(* Logix 5000 project; controller PLC_MCC1201_220AP1 vendor 1 type 14 code 164 rev 35.11; software revision 35.00; part 6 of 25 *)
(* tags used below, declared in another part *)
   B3 : DINT[102];
   HMI_Alarm_Reset : BOOL;   // HMI_Alarm_Reset
   HMI_MAN_CMD_WR : UDT_MAN_CMD_WR;
   LEHR_SPEED : ALIAS FOR N60[1];
   M206_M1_DR : AXIS_CIP_DRIVE;
   M207_M1_DR : AXIS_CIP_DRIVE;
   M208_M1_DR : AXIS_CIP_DRIVE;
   M209_M1_DR : AXIS_CIP_DRIVE;
   M2xx_CONVEYOR : MAC_CONVEYOR[20];
   M2xx_CONVEYOR_IN_MOTION : MAC_CONVEYOR_IN_MOTION[20];
   M2xx_CONVEYOR_OUT_MOTION : MAC_CONVEYOR_OUT_MOTION[20];
   TMP_dDirection : DINT;
   TMP_rAcc : REAL;
   TMP_rDec : REAL;
   TMP_rSpeed : REAL;
   TMP_xAlwaysOFF : BOOL;
   TMP_xRun : BOOL;
(* CommandLogic, continued *)

ROUTINE M206_Conveyor_Motion_Output   (* ladder *)
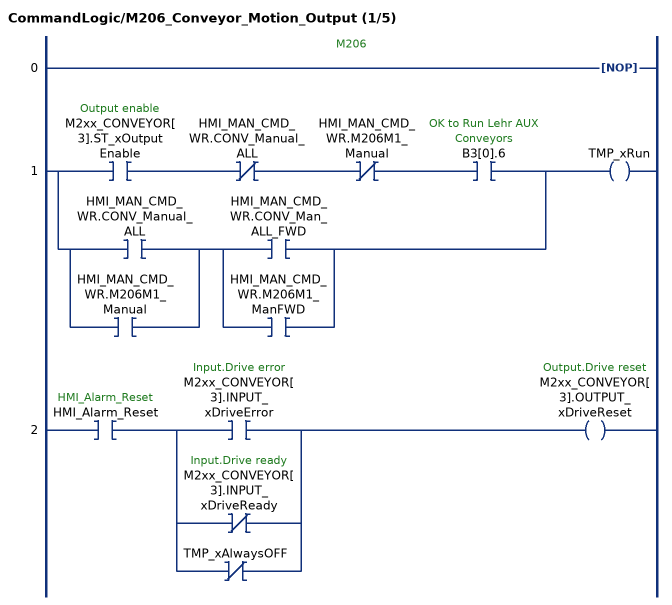
   // M206
   0: NOP();
   1: [XIC(M2xx_CONVEYOR[3].ST_xOutputEnable) XIO(HMI_MAN_CMD_WR.CONV_Manual_ALL) XIO(HMI_MAN_CMD_WR.M206M1_Manual) XIC(B3[0].6) ,[XIC(HMI_MAN_CMD_WR.CONV_Manual_ALL) ,XIC(HMI_MAN_CMD_WR.M206M1_Manual) ] [XIC(HMI_MAN_CMD_WR.CONV_Man_ALL_FWD) ,XIC(HMI_MAN_CMD_WR.M206M1_ManFWD) ] ]OTE(TMP_xRun);
   2: XIC(HMI_Alarm_Reset)[XIC(M2xx_CONVEYOR[3].INPUT_xDriveError) ,XIO(M2xx_CONVEYOR[3].INPUT_xDriveReady) ,XIO(TMP_xAlwaysOFF) ]OTE(M2xx_CONVEYOR[3].OUTPUT_xDriveReset);
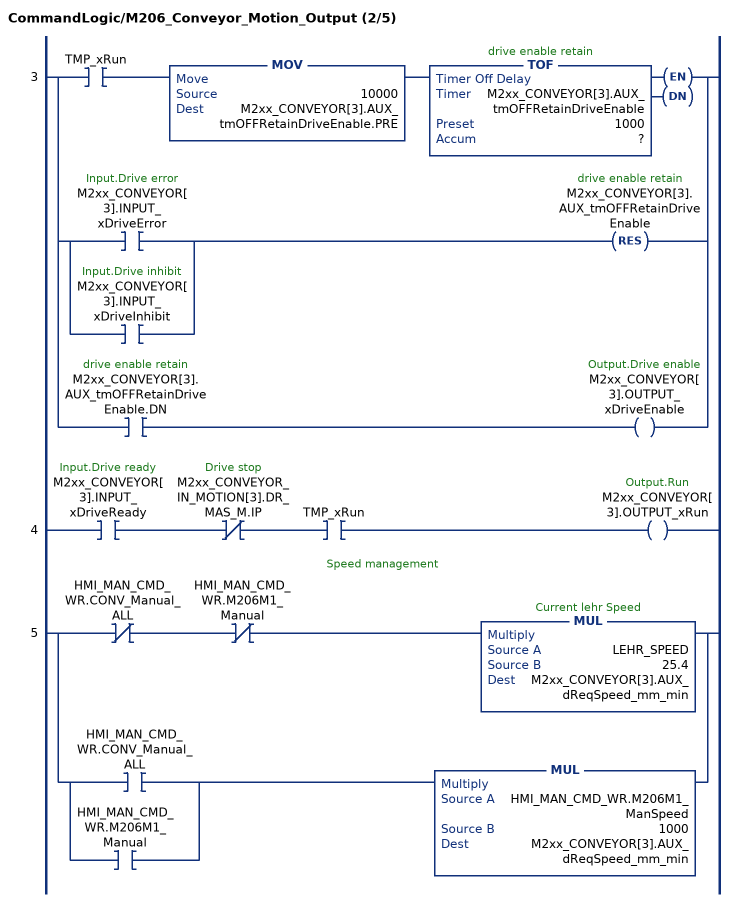
   3: [XIC(TMP_xRun) MOV(10000,M2xx_CONVEYOR[3].AUX_tmOFFRetainDriveEnable.PRE) TOF(M2xx_CONVEYOR[3].AUX_tmOFFRetainDriveEnable,?,?) ,[XIC(M2xx_CONVEYOR[3].INPUT_xDriveError) ,XIC(M2xx_CONVEYOR[3].INPUT_xDriveInhibit) ] RES(M2xx_CONVEYOR[3].AUX_tmOFFRetainDriveEnable) ,XIC(M2xx_CONVEYOR[3].AUX_tmOFFRetainDriveEnable.DN) OTE(M2xx_CONVEYOR[3].OUTPUT_xDriveEnable) ];
   4: XIC(M2xx_CONVEYOR[3].INPUT_xDriveReady)XIO(M2xx_CONVEYOR_IN_MOTION[3].DR_MAS_M.IP)XIC(TMP_xRun)OTE(M2xx_CONVEYOR[3].OUTPUT_xRun);
   // Speed management
   5: [XIO(HMI_MAN_CMD_WR.CONV_Manual_ALL) XIO(HMI_MAN_CMD_WR.M206M1_Manual) MUL(LEHR_SPEED,25.4,M2xx_CONVEYOR[3].AUX_dReqSpeed_mm_min) ,[XIC(HMI_MAN_CMD_WR.CONV_Manual_ALL) ,XIC(HMI_MAN_CMD_WR.M206M1_Manual) ] MUL(HMI_MAN_CMD_WR.M206M1_ManSpeed,1000,M2xx_CONVEYOR[3].AUX_dReqSpeed_mm_min) ];
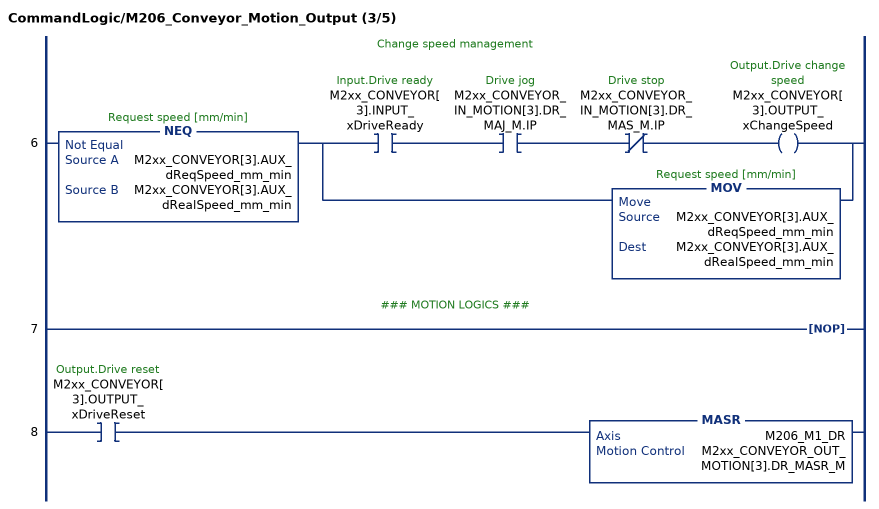
   // Change speed management
   6: NEQ(M2xx_CONVEYOR[3].AUX_dReqSpeed_mm_min,M2xx_CONVEYOR[3].AUX_dRealSpeed_mm_min)[XIC(M2xx_CONVEYOR[3].INPUT_xDriveReady) XIC(M2xx_CONVEYOR_IN_MOTION[3].DR_MAJ_M.IP) XIO(M2xx_CONVEYOR_IN_MOTION[3].DR_MAS_M.IP) OTE(M2xx_CONVEYOR[3].OUTPUT_xChangeSpeed) ,MOV(M2xx_CONVEYOR[3].AUX_dReqSpeed_mm_min,M2xx_CONVEYOR[3].AUX_dRealSpeed_mm_min) ];
   // ### MOTION LOGICS ###
   7: NOP();
   8: XIC(M2xx_CONVEYOR[3].OUTPUT_xDriveReset)MASR(M206_M1_DR,M2xx_CONVEYOR_OUT_MOTION[3].DR_MASR_M);
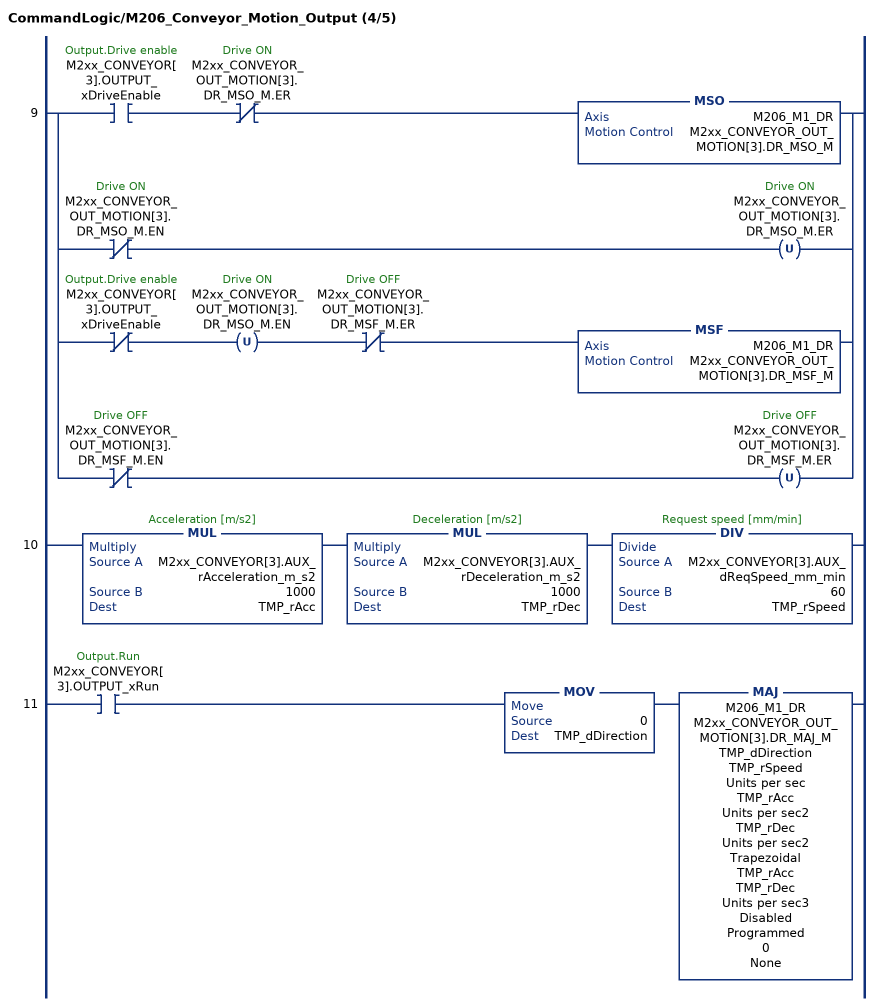
   9: [XIC(M2xx_CONVEYOR[3].OUTPUT_xDriveEnable) XIO(M2xx_CONVEYOR_OUT_MOTION[3].DR_MSO_M.ER) MSO(M206_M1_DR,M2xx_CONVEYOR_OUT_MOTION[3].DR_MSO_M) ,XIO(M2xx_CONVEYOR_OUT_MOTION[3].DR_MSO_M.EN) OTU(M2xx_CONVEYOR_OUT_MOTION[3].DR_MSO_M.ER) ,XIO(M2xx_CONVEYOR[3].OUTPUT_xDriveEnable) OTU(M2xx_CONVEYOR_OUT_MOTION[3].DR_MSO_M.EN) XIO(M2xx_CONVEYOR_OUT_MOTION[3].DR_MSF_M.ER) MSF(M206_M1_DR,M2xx_CONVEYOR_OUT_MOTION[3].DR_MSF_M) ,XIO(M2xx_CONVEYOR_OUT_MOTION[3].DR_MSF_M.EN) OTU(M2xx_CONVEYOR_OUT_MOTION[3].DR_MSF_M.ER) ];
   10: MUL(M2xx_CONVEYOR[3].AUX_rAcceleration_m_s2,1000,TMP_rAcc)MUL(M2xx_CONVEYOR[3].AUX_rDeceleration_m_s2,1000,TMP_rDec)DIV(M2xx_CONVEYOR[3].AUX_dReqSpeed_mm_min,60,TMP_rSpeed);
   11: XIC(M2xx_CONVEYOR[3].OUTPUT_xRun)MOV(0,TMP_dDirection)MAJ(M206_M1_DR,M2xx_CONVEYOR_OUT_MOTION[3].DR_MAJ_M,TMP_dDirection,TMP_rSpeed,Units per sec,TMP_rAcc,Units per sec2,TMP_rDec,Units per sec2,Trapezoidal,TMP_rAcc,TMP_rDec,Units per sec3,Disabled,Programmed,0,None);
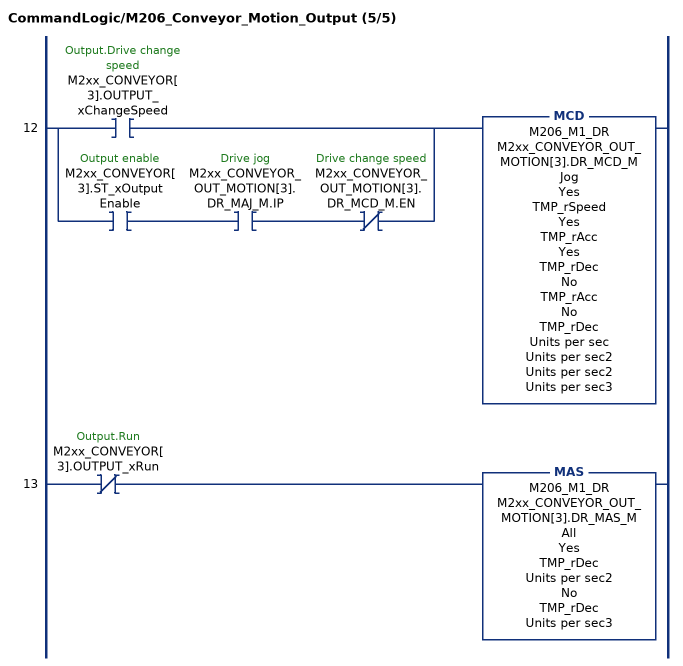
   12: [XIC(M2xx_CONVEYOR[3].OUTPUT_xChangeSpeed) ,XIC(M2xx_CONVEYOR[3].ST_xOutputEnable) XIC(M2xx_CONVEYOR_OUT_MOTION[3].DR_MAJ_M.IP) XIO(M2xx_CONVEYOR_OUT_MOTION[3].DR_MCD_M.EN) ]MCD(M206_M1_DR,M2xx_CONVEYOR_OUT_MOTION[3].DR_MCD_M,Jog,Yes,TMP_rSpeed,Yes,TMP_rAcc,Yes,TMP_rDec,No,TMP_rAcc,No,TMP_rDec,Units per sec,Units per sec2,Units per sec2,Units per sec3);
   13: XIO(M2xx_CONVEYOR[3].OUTPUT_xRun)MAS(M206_M1_DR,M2xx_CONVEYOR_OUT_MOTION[3].DR_MAS_M,All,Yes,TMP_rDec,Units per sec2,No,TMP_rDec,Units per sec3);
END_ROUTINE

ROUTINE M207_Conveyor_Motion_Output   (* ladder *)
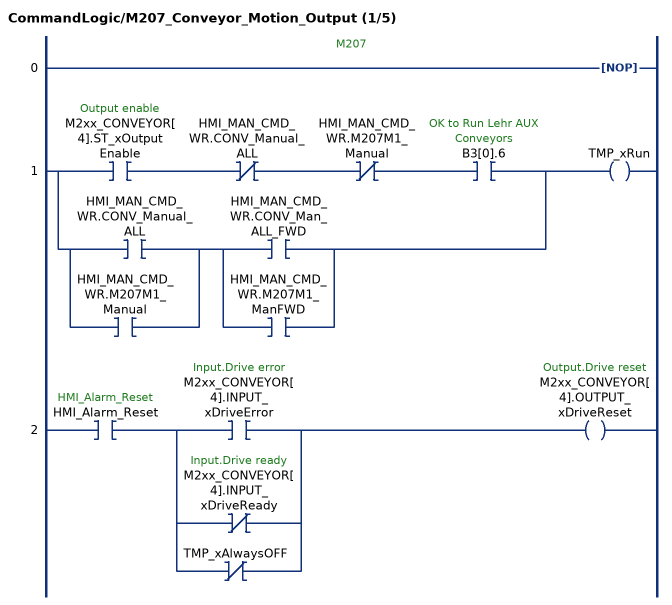
   // M207
   0: NOP();
   1: [XIC(M2xx_CONVEYOR[4].ST_xOutputEnable) XIO(HMI_MAN_CMD_WR.CONV_Manual_ALL) XIO(HMI_MAN_CMD_WR.M207M1_Manual) XIC(B3[0].6) ,[XIC(HMI_MAN_CMD_WR.CONV_Manual_ALL) ,XIC(HMI_MAN_CMD_WR.M207M1_Manual) ] [XIC(HMI_MAN_CMD_WR.CONV_Man_ALL_FWD) ,XIC(HMI_MAN_CMD_WR.M207M1_ManFWD) ] ]OTE(TMP_xRun);
   2: XIC(HMI_Alarm_Reset)[XIC(M2xx_CONVEYOR[4].INPUT_xDriveError) ,XIO(M2xx_CONVEYOR[4].INPUT_xDriveReady) ,XIO(TMP_xAlwaysOFF) ]OTE(M2xx_CONVEYOR[4].OUTPUT_xDriveReset);
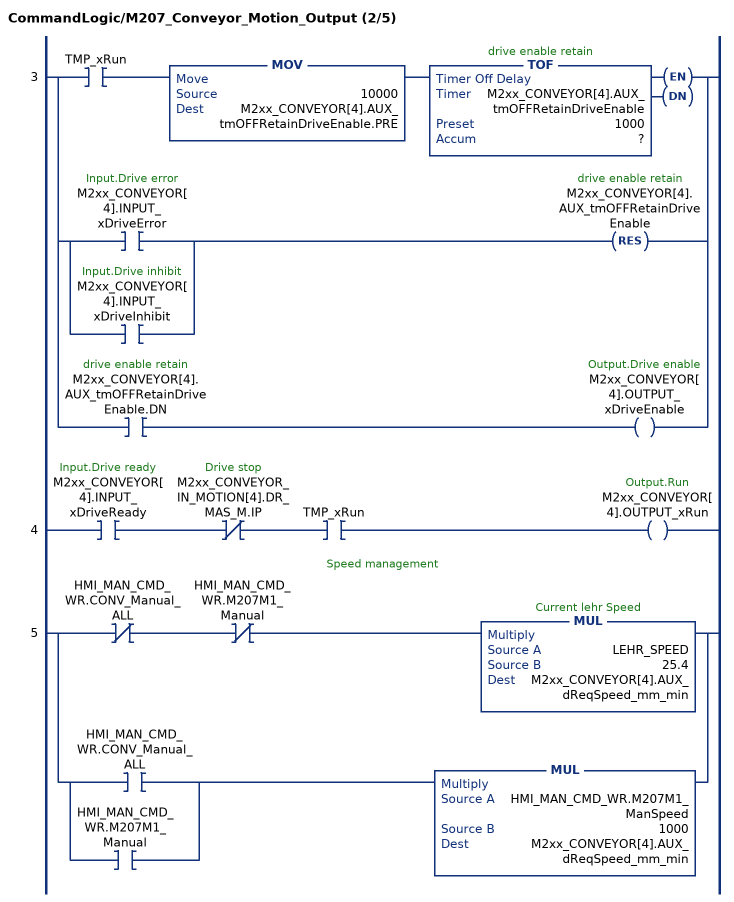
   3: [XIC(TMP_xRun) MOV(10000,M2xx_CONVEYOR[4].AUX_tmOFFRetainDriveEnable.PRE) TOF(M2xx_CONVEYOR[4].AUX_tmOFFRetainDriveEnable,?,?) ,[XIC(M2xx_CONVEYOR[4].INPUT_xDriveError) ,XIC(M2xx_CONVEYOR[4].INPUT_xDriveInhibit) ] RES(M2xx_CONVEYOR[4].AUX_tmOFFRetainDriveEnable) ,XIC(M2xx_CONVEYOR[4].AUX_tmOFFRetainDriveEnable.DN) OTE(M2xx_CONVEYOR[4].OUTPUT_xDriveEnable) ];
   4: XIC(M2xx_CONVEYOR[4].INPUT_xDriveReady)XIO(M2xx_CONVEYOR_IN_MOTION[4].DR_MAS_M.IP)XIC(TMP_xRun)OTE(M2xx_CONVEYOR[4].OUTPUT_xRun);
   // Speed management
   5: [XIO(HMI_MAN_CMD_WR.CONV_Manual_ALL) XIO(HMI_MAN_CMD_WR.M207M1_Manual) MUL(LEHR_SPEED,25.4,M2xx_CONVEYOR[4].AUX_dReqSpeed_mm_min) ,[XIC(HMI_MAN_CMD_WR.CONV_Manual_ALL) ,XIC(HMI_MAN_CMD_WR.M207M1_Manual) ] MUL(HMI_MAN_CMD_WR.M207M1_ManSpeed,1000,M2xx_CONVEYOR[4].AUX_dReqSpeed_mm_min) ];
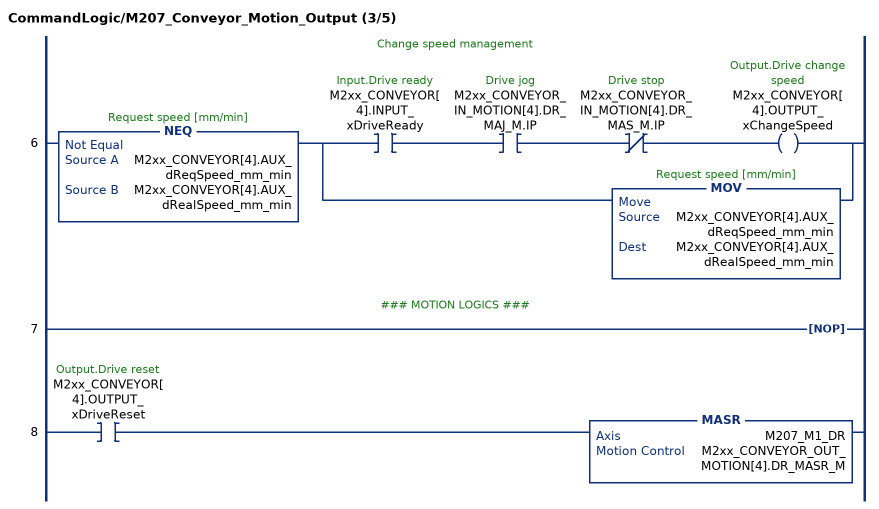
   // Change speed management
   6: NEQ(M2xx_CONVEYOR[4].AUX_dReqSpeed_mm_min,M2xx_CONVEYOR[4].AUX_dRealSpeed_mm_min)[XIC(M2xx_CONVEYOR[4].INPUT_xDriveReady) XIC(M2xx_CONVEYOR_IN_MOTION[4].DR_MAJ_M.IP) XIO(M2xx_CONVEYOR_IN_MOTION[4].DR_MAS_M.IP) OTE(M2xx_CONVEYOR[4].OUTPUT_xChangeSpeed) ,MOV(M2xx_CONVEYOR[4].AUX_dReqSpeed_mm_min,M2xx_CONVEYOR[4].AUX_dRealSpeed_mm_min) ];
   // ### MOTION LOGICS ###
   7: NOP();
   8: XIC(M2xx_CONVEYOR[4].OUTPUT_xDriveReset)MASR(M207_M1_DR,M2xx_CONVEYOR_OUT_MOTION[4].DR_MASR_M);
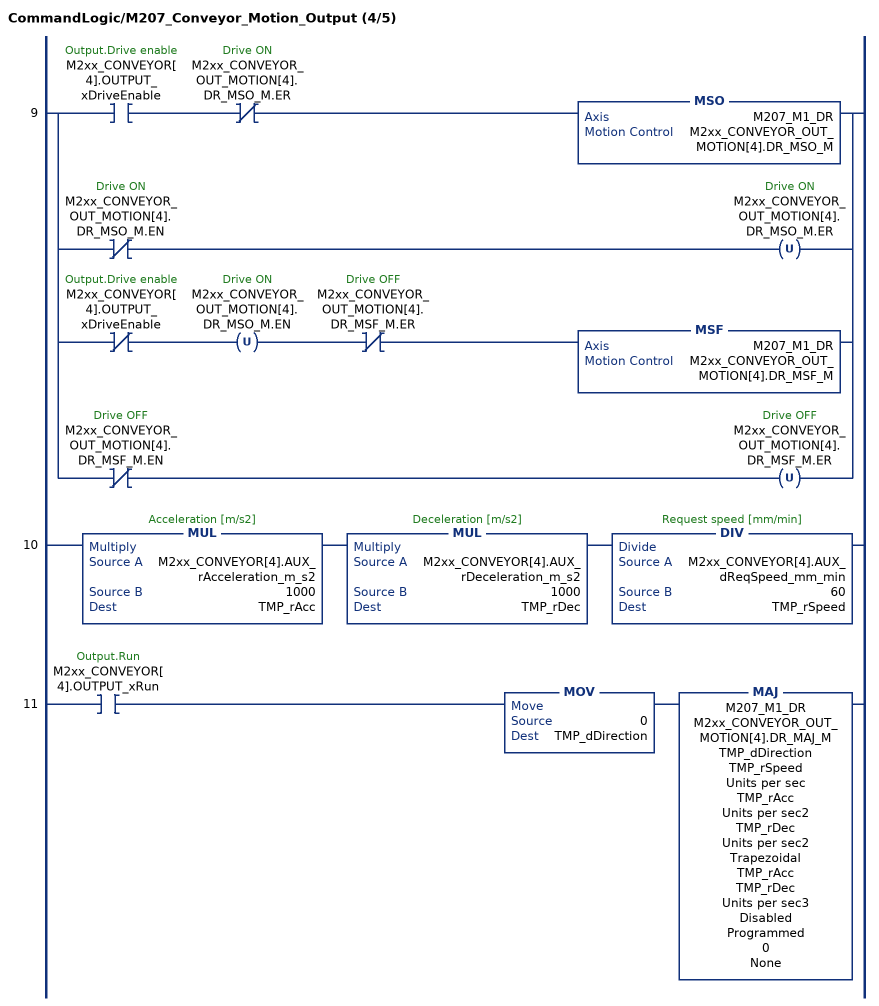
   9: [XIC(M2xx_CONVEYOR[4].OUTPUT_xDriveEnable) XIO(M2xx_CONVEYOR_OUT_MOTION[4].DR_MSO_M.ER) MSO(M207_M1_DR,M2xx_CONVEYOR_OUT_MOTION[4].DR_MSO_M) ,XIO(M2xx_CONVEYOR_OUT_MOTION[4].DR_MSO_M.EN) OTU(M2xx_CONVEYOR_OUT_MOTION[4].DR_MSO_M.ER) ,XIO(M2xx_CONVEYOR[4].OUTPUT_xDriveEnable) OTU(M2xx_CONVEYOR_OUT_MOTION[4].DR_MSO_M.EN) XIO(M2xx_CONVEYOR_OUT_MOTION[4].DR_MSF_M.ER) MSF(M207_M1_DR,M2xx_CONVEYOR_OUT_MOTION[4].DR_MSF_M) ,XIO(M2xx_CONVEYOR_OUT_MOTION[4].DR_MSF_M.EN) OTU(M2xx_CONVEYOR_OUT_MOTION[4].DR_MSF_M.ER) ];
   10: MUL(M2xx_CONVEYOR[4].AUX_rAcceleration_m_s2,1000,TMP_rAcc)MUL(M2xx_CONVEYOR[4].AUX_rDeceleration_m_s2,1000,TMP_rDec)DIV(M2xx_CONVEYOR[4].AUX_dReqSpeed_mm_min,60,TMP_rSpeed);
   11: XIC(M2xx_CONVEYOR[4].OUTPUT_xRun)MOV(0,TMP_dDirection)MAJ(M207_M1_DR,M2xx_CONVEYOR_OUT_MOTION[4].DR_MAJ_M,TMP_dDirection,TMP_rSpeed,Units per sec,TMP_rAcc,Units per sec2,TMP_rDec,Units per sec2,Trapezoidal,TMP_rAcc,TMP_rDec,Units per sec3,Disabled,Programmed,0,None);
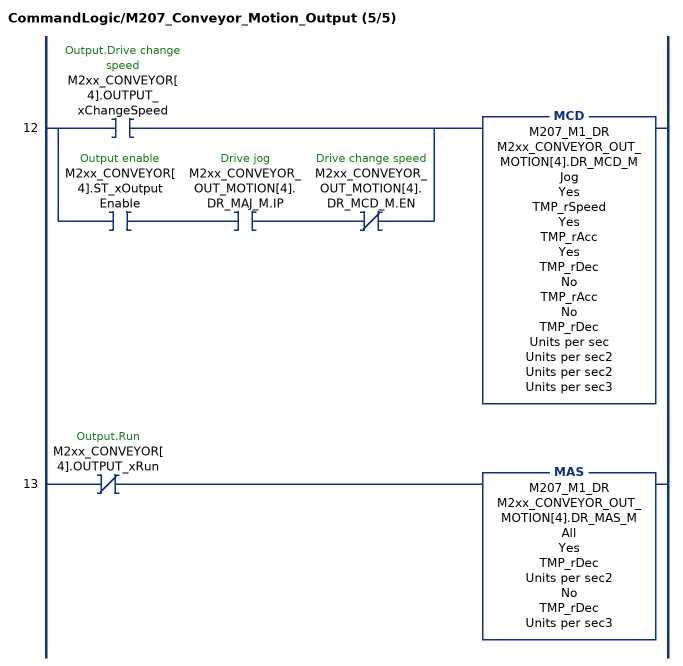
   12: [XIC(M2xx_CONVEYOR[4].OUTPUT_xChangeSpeed) ,XIC(M2xx_CONVEYOR[4].ST_xOutputEnable) XIC(M2xx_CONVEYOR_OUT_MOTION[4].DR_MAJ_M.IP) XIO(M2xx_CONVEYOR_OUT_MOTION[4].DR_MCD_M.EN) ]MCD(M207_M1_DR,M2xx_CONVEYOR_OUT_MOTION[4].DR_MCD_M,Jog,Yes,TMP_rSpeed,Yes,TMP_rAcc,Yes,TMP_rDec,No,TMP_rAcc,No,TMP_rDec,Units per sec,Units per sec2,Units per sec2,Units per sec3);
   13: XIO(M2xx_CONVEYOR[4].OUTPUT_xRun)MAS(M207_M1_DR,M2xx_CONVEYOR_OUT_MOTION[4].DR_MAS_M,All,Yes,TMP_rDec,Units per sec2,No,TMP_rDec,Units per sec3);
END_ROUTINE

ROUTINE M208_Conveyor_Motion_Output   (* ladder *)
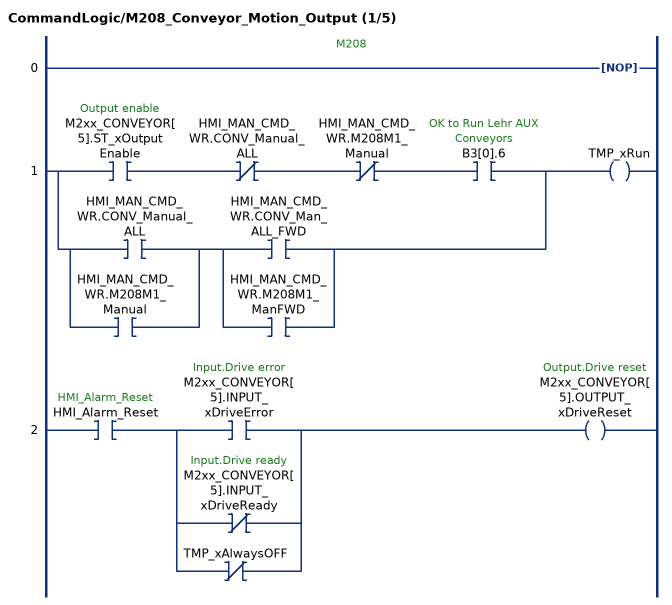
   // M208
   0: NOP();
   1: [XIC(M2xx_CONVEYOR[5].ST_xOutputEnable) XIO(HMI_MAN_CMD_WR.CONV_Manual_ALL) XIO(HMI_MAN_CMD_WR.M208M1_Manual) XIC(B3[0].6) ,[XIC(HMI_MAN_CMD_WR.CONV_Manual_ALL) ,XIC(HMI_MAN_CMD_WR.M208M1_Manual) ] [XIC(HMI_MAN_CMD_WR.CONV_Man_ALL_FWD) ,XIC(HMI_MAN_CMD_WR.M208M1_ManFWD) ] ]OTE(TMP_xRun);
   2: XIC(HMI_Alarm_Reset)[XIC(M2xx_CONVEYOR[5].INPUT_xDriveError) ,XIO(M2xx_CONVEYOR[5].INPUT_xDriveReady) ,XIO(TMP_xAlwaysOFF) ]OTE(M2xx_CONVEYOR[5].OUTPUT_xDriveReset);
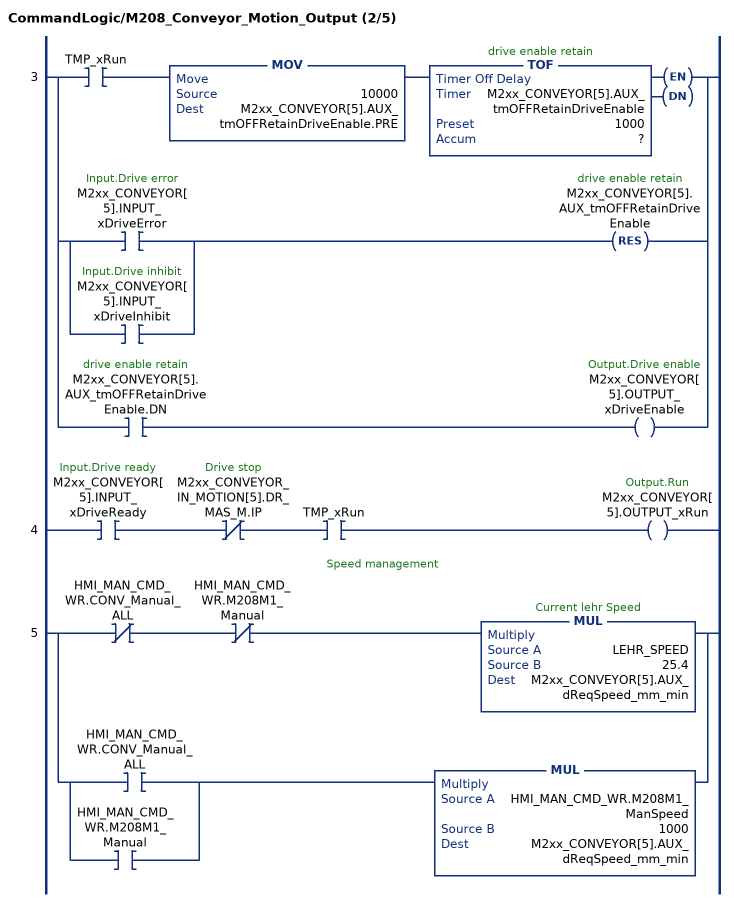
   3: [XIC(TMP_xRun) MOV(10000,M2xx_CONVEYOR[5].AUX_tmOFFRetainDriveEnable.PRE) TOF(M2xx_CONVEYOR[5].AUX_tmOFFRetainDriveEnable,?,?) ,[XIC(M2xx_CONVEYOR[5].INPUT_xDriveError) ,XIC(M2xx_CONVEYOR[5].INPUT_xDriveInhibit) ] RES(M2xx_CONVEYOR[5].AUX_tmOFFRetainDriveEnable) ,XIC(M2xx_CONVEYOR[5].AUX_tmOFFRetainDriveEnable.DN) OTE(M2xx_CONVEYOR[5].OUTPUT_xDriveEnable) ];
   4: XIC(M2xx_CONVEYOR[5].INPUT_xDriveReady)XIO(M2xx_CONVEYOR_IN_MOTION[5].DR_MAS_M.IP)XIC(TMP_xRun)OTE(M2xx_CONVEYOR[5].OUTPUT_xRun);
   // Speed management
   5: [XIO(HMI_MAN_CMD_WR.CONV_Manual_ALL) XIO(HMI_MAN_CMD_WR.M208M1_Manual) MUL(LEHR_SPEED,25.4,M2xx_CONVEYOR[5].AUX_dReqSpeed_mm_min) ,[XIC(HMI_MAN_CMD_WR.CONV_Manual_ALL) ,XIC(HMI_MAN_CMD_WR.M208M1_Manual) ] MUL(HMI_MAN_CMD_WR.M208M1_ManSpeed,1000,M2xx_CONVEYOR[5].AUX_dReqSpeed_mm_min) ];
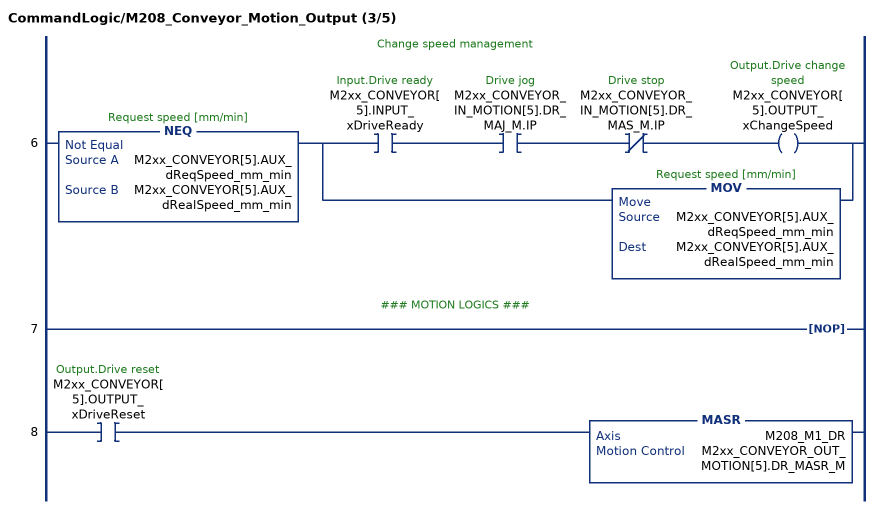
   // Change speed management
   6: NEQ(M2xx_CONVEYOR[5].AUX_dReqSpeed_mm_min,M2xx_CONVEYOR[5].AUX_dRealSpeed_mm_min)[XIC(M2xx_CONVEYOR[5].INPUT_xDriveReady) XIC(M2xx_CONVEYOR_IN_MOTION[5].DR_MAJ_M.IP) XIO(M2xx_CONVEYOR_IN_MOTION[5].DR_MAS_M.IP) OTE(M2xx_CONVEYOR[5].OUTPUT_xChangeSpeed) ,MOV(M2xx_CONVEYOR[5].AUX_dReqSpeed_mm_min,M2xx_CONVEYOR[5].AUX_dRealSpeed_mm_min) ];
   // ### MOTION LOGICS ###
   7: NOP();
   8: XIC(M2xx_CONVEYOR[5].OUTPUT_xDriveReset)MASR(M208_M1_DR,M2xx_CONVEYOR_OUT_MOTION[5].DR_MASR_M);
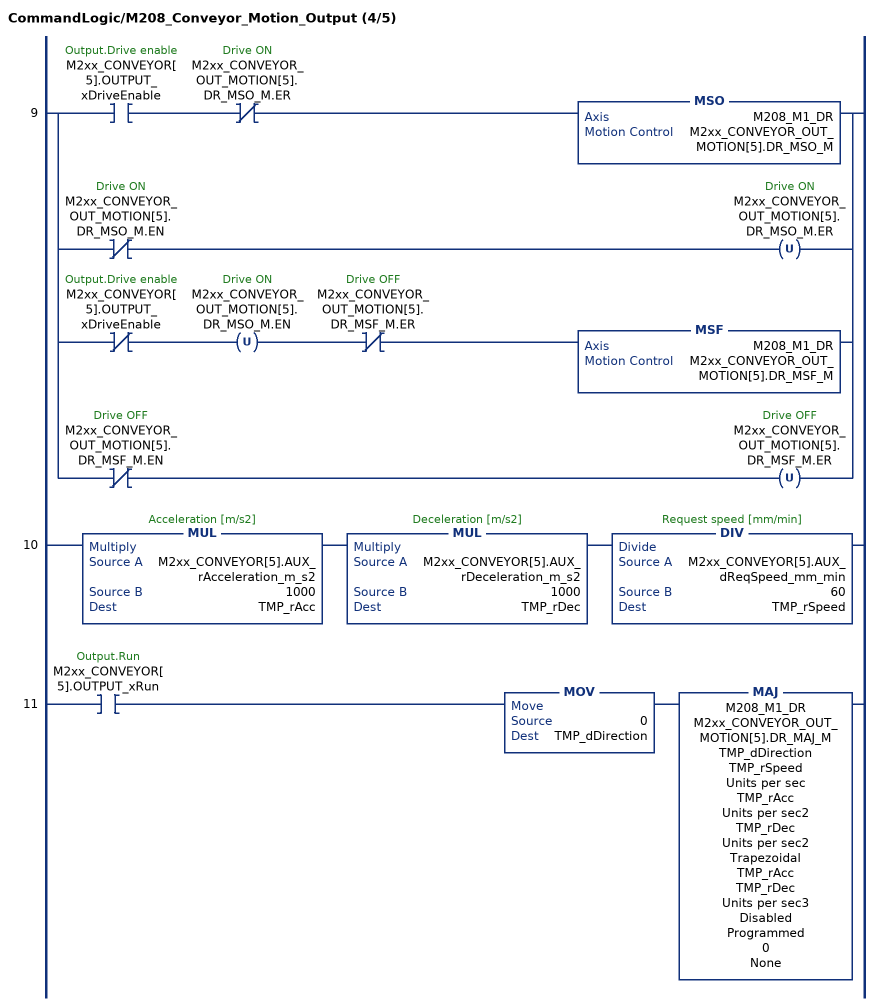
   9: [XIC(M2xx_CONVEYOR[5].OUTPUT_xDriveEnable) XIO(M2xx_CONVEYOR_OUT_MOTION[5].DR_MSO_M.ER) MSO(M208_M1_DR,M2xx_CONVEYOR_OUT_MOTION[5].DR_MSO_M) ,XIO(M2xx_CONVEYOR_OUT_MOTION[5].DR_MSO_M.EN) OTU(M2xx_CONVEYOR_OUT_MOTION[5].DR_MSO_M.ER) ,XIO(M2xx_CONVEYOR[5].OUTPUT_xDriveEnable) OTU(M2xx_CONVEYOR_OUT_MOTION[5].DR_MSO_M.EN) XIO(M2xx_CONVEYOR_OUT_MOTION[5].DR_MSF_M.ER) MSF(M208_M1_DR,M2xx_CONVEYOR_OUT_MOTION[5].DR_MSF_M) ,XIO(M2xx_CONVEYOR_OUT_MOTION[5].DR_MSF_M.EN) OTU(M2xx_CONVEYOR_OUT_MOTION[5].DR_MSF_M.ER) ];
   10: MUL(M2xx_CONVEYOR[5].AUX_rAcceleration_m_s2,1000,TMP_rAcc)MUL(M2xx_CONVEYOR[5].AUX_rDeceleration_m_s2,1000,TMP_rDec)DIV(M2xx_CONVEYOR[5].AUX_dReqSpeed_mm_min,60,TMP_rSpeed);
   11: XIC(M2xx_CONVEYOR[5].OUTPUT_xRun)MOV(0,TMP_dDirection)MAJ(M208_M1_DR,M2xx_CONVEYOR_OUT_MOTION[5].DR_MAJ_M,TMP_dDirection,TMP_rSpeed,Units per sec,TMP_rAcc,Units per sec2,TMP_rDec,Units per sec2,Trapezoidal,TMP_rAcc,TMP_rDec,Units per sec3,Disabled,Programmed,0,None);
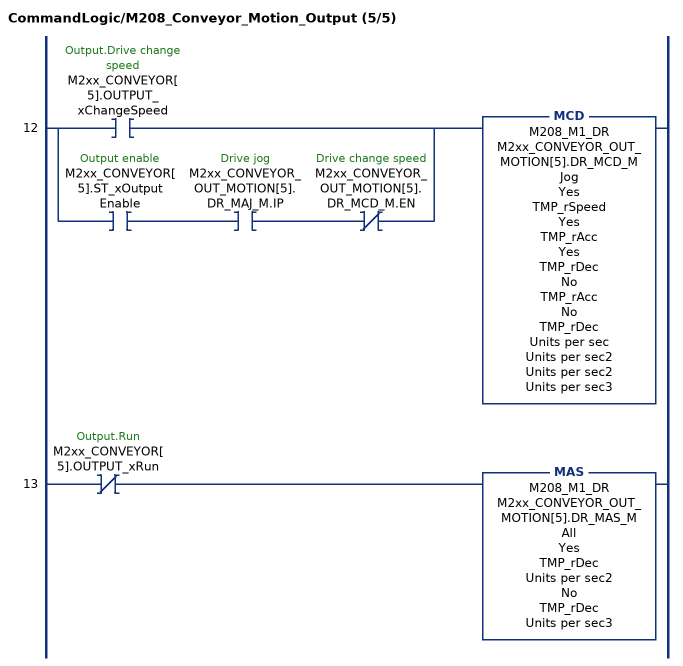
   12: [XIC(M2xx_CONVEYOR[5].OUTPUT_xChangeSpeed) ,XIC(M2xx_CONVEYOR[5].ST_xOutputEnable) XIC(M2xx_CONVEYOR_OUT_MOTION[5].DR_MAJ_M.IP) XIO(M2xx_CONVEYOR_OUT_MOTION[5].DR_MCD_M.EN) ]MCD(M208_M1_DR,M2xx_CONVEYOR_OUT_MOTION[5].DR_MCD_M,Jog,Yes,TMP_rSpeed,Yes,TMP_rAcc,Yes,TMP_rDec,No,TMP_rAcc,No,TMP_rDec,Units per sec,Units per sec2,Units per sec2,Units per sec3);
   13: XIO(M2xx_CONVEYOR[5].OUTPUT_xRun)MAS(M208_M1_DR,M2xx_CONVEYOR_OUT_MOTION[5].DR_MAS_M,All,Yes,TMP_rDec,Units per sec2,No,TMP_rDec,Units per sec3);
END_ROUTINE

ROUTINE M209_Conveyor_Motion_Output   (* ladder *)
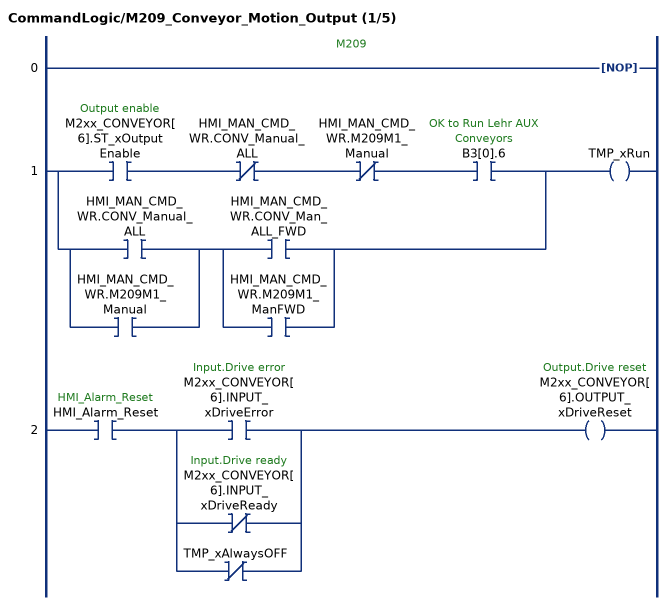
   // M209
   0: NOP();
   1: [XIC(M2xx_CONVEYOR[6].ST_xOutputEnable) XIO(HMI_MAN_CMD_WR.CONV_Manual_ALL) XIO(HMI_MAN_CMD_WR.M209M1_Manual) XIC(B3[0].6) ,[XIC(HMI_MAN_CMD_WR.CONV_Manual_ALL) ,XIC(HMI_MAN_CMD_WR.M209M1_Manual) ] [XIC(HMI_MAN_CMD_WR.CONV_Man_ALL_FWD) ,XIC(HMI_MAN_CMD_WR.M209M1_ManFWD) ] ]OTE(TMP_xRun);
   2: XIC(HMI_Alarm_Reset)[XIC(M2xx_CONVEYOR[6].INPUT_xDriveError) ,XIO(M2xx_CONVEYOR[6].INPUT_xDriveReady) ,XIO(TMP_xAlwaysOFF) ]OTE(M2xx_CONVEYOR[6].OUTPUT_xDriveReset);
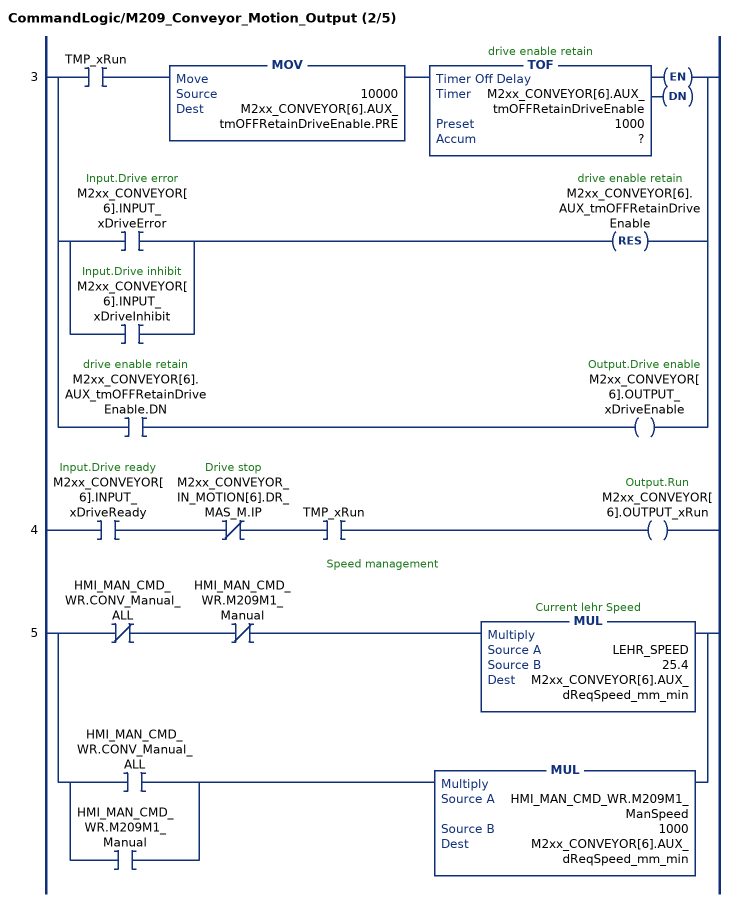
   3: [XIC(TMP_xRun) MOV(10000,M2xx_CONVEYOR[6].AUX_tmOFFRetainDriveEnable.PRE) TOF(M2xx_CONVEYOR[6].AUX_tmOFFRetainDriveEnable,?,?) ,[XIC(M2xx_CONVEYOR[6].INPUT_xDriveError) ,XIC(M2xx_CONVEYOR[6].INPUT_xDriveInhibit) ] RES(M2xx_CONVEYOR[6].AUX_tmOFFRetainDriveEnable) ,XIC(M2xx_CONVEYOR[6].AUX_tmOFFRetainDriveEnable.DN) OTE(M2xx_CONVEYOR[6].OUTPUT_xDriveEnable) ];
   4: XIC(M2xx_CONVEYOR[6].INPUT_xDriveReady)XIO(M2xx_CONVEYOR_IN_MOTION[6].DR_MAS_M.IP)XIC(TMP_xRun)OTE(M2xx_CONVEYOR[6].OUTPUT_xRun);
   // Speed management
   5: [XIO(HMI_MAN_CMD_WR.CONV_Manual_ALL) XIO(HMI_MAN_CMD_WR.M209M1_Manual) MUL(LEHR_SPEED,25.4,M2xx_CONVEYOR[6].AUX_dReqSpeed_mm_min) ,[XIC(HMI_MAN_CMD_WR.CONV_Manual_ALL) ,XIC(HMI_MAN_CMD_WR.M209M1_Manual) ] MUL(HMI_MAN_CMD_WR.M209M1_ManSpeed,1000,M2xx_CONVEYOR[6].AUX_dReqSpeed_mm_min) ];
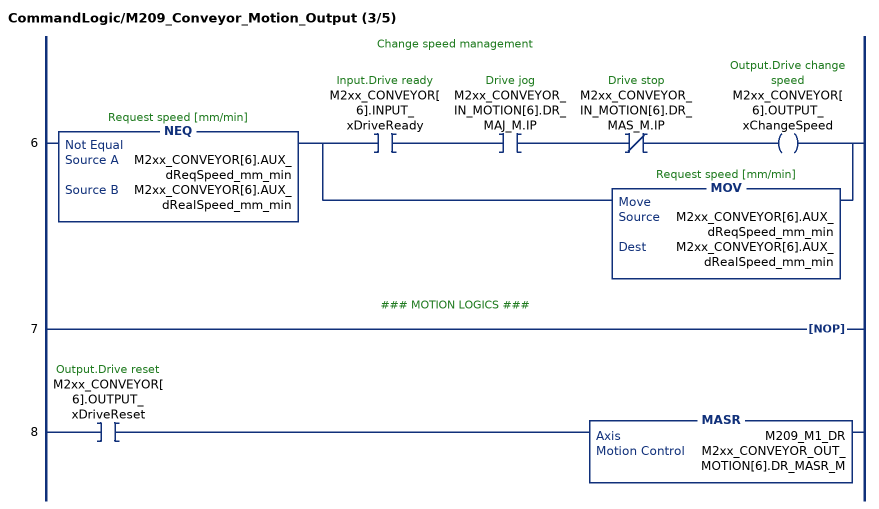
   // Change speed management
   6: NEQ(M2xx_CONVEYOR[6].AUX_dReqSpeed_mm_min,M2xx_CONVEYOR[6].AUX_dRealSpeed_mm_min)[XIC(M2xx_CONVEYOR[6].INPUT_xDriveReady) XIC(M2xx_CONVEYOR_IN_MOTION[6].DR_MAJ_M.IP) XIO(M2xx_CONVEYOR_IN_MOTION[6].DR_MAS_M.IP) OTE(M2xx_CONVEYOR[6].OUTPUT_xChangeSpeed) ,MOV(M2xx_CONVEYOR[6].AUX_dReqSpeed_mm_min,M2xx_CONVEYOR[6].AUX_dRealSpeed_mm_min) ];
   // ### MOTION LOGICS ###
   7: NOP();
   8: XIC(M2xx_CONVEYOR[6].OUTPUT_xDriveReset)MASR(M209_M1_DR,M2xx_CONVEYOR_OUT_MOTION[6].DR_MASR_M);
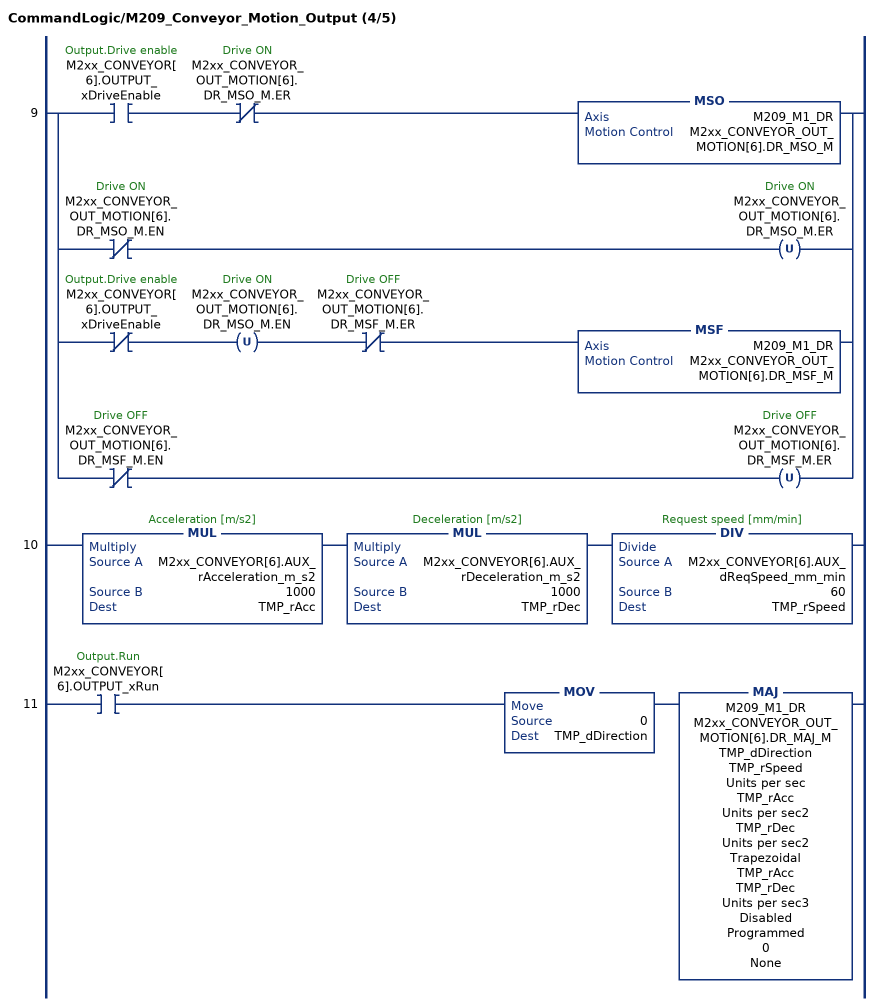
   9: [XIC(M2xx_CONVEYOR[6].OUTPUT_xDriveEnable) XIO(M2xx_CONVEYOR_OUT_MOTION[6].DR_MSO_M.ER) MSO(M209_M1_DR,M2xx_CONVEYOR_OUT_MOTION[6].DR_MSO_M) ,XIO(M2xx_CONVEYOR_OUT_MOTION[6].DR_MSO_M.EN) OTU(M2xx_CONVEYOR_OUT_MOTION[6].DR_MSO_M.ER) ,XIO(M2xx_CONVEYOR[6].OUTPUT_xDriveEnable) OTU(M2xx_CONVEYOR_OUT_MOTION[6].DR_MSO_M.EN) XIO(M2xx_CONVEYOR_OUT_MOTION[6].DR_MSF_M.ER) MSF(M209_M1_DR,M2xx_CONVEYOR_OUT_MOTION[6].DR_MSF_M) ,XIO(M2xx_CONVEYOR_OUT_MOTION[6].DR_MSF_M.EN) OTU(M2xx_CONVEYOR_OUT_MOTION[6].DR_MSF_M.ER) ];
   10: MUL(M2xx_CONVEYOR[6].AUX_rAcceleration_m_s2,1000,TMP_rAcc)MUL(M2xx_CONVEYOR[6].AUX_rDeceleration_m_s2,1000,TMP_rDec)DIV(M2xx_CONVEYOR[6].AUX_dReqSpeed_mm_min,60,TMP_rSpeed);
   11: XIC(M2xx_CONVEYOR[6].OUTPUT_xRun)MOV(0,TMP_dDirection)MAJ(M209_M1_DR,M2xx_CONVEYOR_OUT_MOTION[6].DR_MAJ_M,TMP_dDirection,TMP_rSpeed,Units per sec,TMP_rAcc,Units per sec2,TMP_rDec,Units per sec2,Trapezoidal,TMP_rAcc,TMP_rDec,Units per sec3,Disabled,Programmed,0,None);
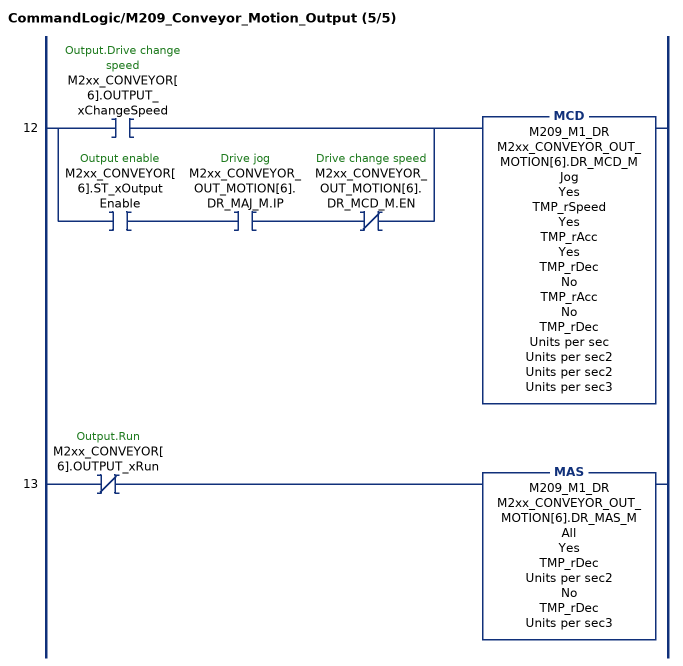
   12: [XIC(M2xx_CONVEYOR[6].OUTPUT_xChangeSpeed) ,XIC(M2xx_CONVEYOR[6].ST_xOutputEnable) XIC(M2xx_CONVEYOR_OUT_MOTION[6].DR_MAJ_M.IP) XIO(M2xx_CONVEYOR_OUT_MOTION[6].DR_MCD_M.EN) ]MCD(M209_M1_DR,M2xx_CONVEYOR_OUT_MOTION[6].DR_MCD_M,Jog,Yes,TMP_rSpeed,Yes,TMP_rAcc,Yes,TMP_rDec,No,TMP_rAcc,No,TMP_rDec,Units per sec,Units per sec2,Units per sec2,Units per sec3);
   13: XIO(M2xx_CONVEYOR[6].OUTPUT_xRun)MAS(M209_M1_DR,M2xx_CONVEYOR_OUT_MOTION[6].DR_MAS_M,All,Yes,TMP_rDec,Units per sec2,No,TMP_rDec,Units per sec3);
END_ROUTINE
